
             IF #statPrevOutputValue >= #inputValue
             THEN
               IF #setPosDownRateLim = 0.0
               THEN
                 // set notification for down rate limit in pos range              
                 #tempPosDown := TRUE;
                 IF #inputValue >= 0.0
                 THEN
                   #tempOutv := #inputValue;
                 ELSE
                   #tempOutv := 0.0;
                 END_IF;
               ELSE
                 IF #inputValue >= 0.0
                 THEN
                   // limited rate of change
                   #tempVar := #statPrevOutputValue - #setPosDownRateLim * #tempCycleReal;
                   IF #inputValue < #tempVar
                   THEN
                     // set notification for up rate limit in pos range                  
                     #tempPosDown := TRUE;
                     #tempOutv := #tempVar;
                   END_IF;
                 ELSE  // changeover between pos. and neg. range
                   // period till zero-crossing
                   #tempVar := #statPrevOutputValue / #setPosDownRateLim;

                   IF #tempVar <= #tempCycleReal
                   THEN
                     // limited rate of change
                     #tempVar := - (#tempCycleReal - #tempVar) * #setNegUpRateLim;

                     IF #inputValue < #tempVar
                     THEN
                       // set notification for rate limit
                       #tempPosDown := False;
                       #tempNegUp := TRUE;
                       #tempOutv := #tempVar;
                     END_IF;
                   ELSE
                     // set notification for rate limit
                     #tempPosDown := TRUE;
                     #tempNegUp := FALSE;
                     #tempOutv := #statPrevOutputValue - #tempCycleReal * #setPosDownRateLim;
                   END_IF;
                 END_IF;
               END_IF;
             END_IF;
           END_IF;
         END_IF;
       END_IF;

       // high/low level limitation
       IF #tempOutv >= #setHighLim
       THEN
         #tempHighLim := TRUE;
         IF NOT #statManOp
         THEN
           #tempOutv := #setHighLim;
           // correct up rate limit notification                
           IF #tempOutv - #statPrevOutputValue < #setPosUpRateLim * #tempCycleReal
           THEN
             #tempPosUp := FALSE;
           END_IF;
         END_IF;
       ELSE
         IF #tempOutv <= #setLowLim
         THEN
           #tempLowLim := TRUE;
           IF NOT #statManOp
           THEN
             #tempOutv := #setLowLim;
             // correct up rate limit notification  
             IF #statPrevOutputValue - #tempOutv < #setNegUpRateLim * #tempCycleReal
             THEN
               #tempNegUp := FALSE;
             END_IF;
           END_IF;
         ELSE
           // reset manual mode flag when tempOutv between upper and lower limit        
           #statManOp := FALSE;
         END_IF;
       END_IF;
     END_IF;
   END_IF;


   // update output parameters
   #outputValue := #tempOutv;    // output
   #statPrevOutputValue := #tempOutv;
   #posUpRateLim := #tempPosUp;
   #posDownRateLim := #tempPosDown;
   #negUpRateLim := #tempNegUp;
   #negDownRateLim := #tempNegDown;
   #highLim := #tempHighLim;
   #lowLim := #tempLowLim;
END_FUNCTION_BLOCK

// folder: Phisical_functions/LGF/8 Technology operations/LGF_NonLin

FUNCTION_BLOCK "LGF_NonLin"   // FB10035, SCL
{ S7_Optimized_Access := 'TRUE' }
VERSION : 2.0
   VAR_INPUT
      inputValue : Real;   // Input value
      defaultOutValue : Real;   // Default output value
      onDefaultOutValue : Bool;   // Default output ON: outputValue = defaultOutputValue
      track : Bool;   // Tracking output ON: outputValue = inputValue
      reset : Bool;   // Complete Restart of function block (outputValue = 0.0)
   END_VAR
   VAR_OUTPUT
      outputValue : Real;   // Output value
   END_VAR
   VAR_IN_OUT
      setpoints : Array[*] of "LGF_typeNonLinSetpoints";   // Setpoint table of polynom
   END_VAR
   VAR
      statIndex : Int;   // Index of setpoint table
   END_VAR
   VAR_TEMP
      tempEndOfSearch : Bool;   // End of search algorithm
      tempInputValueStart : Real;   // Actual setpoint - Input value - Low level
      tempInputValueEnd : Real;   // Actual setpoint - Input value - High level
      tempOutputValueStart : Real;   // Actual setpoint - Output value - Low level
      tempOutputValueEnd : Real;   // Actual setpoint - Output value - High level
      tempFactor : Real;   // Gradient of the straight line
      tempLowerBound : Int;   // -
      tempUpperBound : Int;   // -
   END_VAR
BEGIN
   //=============================================================================
   // SIEMENS AG
   // (c)Copyright 2017
   //-----------------------------------------------------------------------------
   // Library:      LGF(Library General Functions)
   // System:       CPU1212C DC/DC/DC FW:V4.2
   // Engineering:  TIA Portal V14 Update 1
   // Restrictions: -
   // Requirements: PLC (S7-1200 FW: 4.2 / S7-1500 FW: 2.0) or higher
   //-----------------------------------------------------------------------------
   // Change log table:
   // Version date         In charge / Changes applied
   // 01.00.00 04.01.2017  Siemens Industry Online Support
   //                      First released version
   // 01.00.01 17.08.2018  Siemens Industry Online Support
   //                      Upgrade: TIA V15 Update 2
   // 01.00.02 23.11.2018  Siemens Industry Online Support
   //                      Upgrade: TIA V15.1
   //=============================================================================

   //Call "LOWER_BOUND" and "UPPER_BOUND" for the setpoints
   #tempLowerBound := DINT_TO_INT(LOWER_BOUND(ARR := #setpoints, DIM := 1));
   #tempUpperBound := DINT_TO_INT(UPPER_BOUND(ARR := #setpoints, DIM := 1));

   //Check index value
   IF (#statIndex < #tempLowerBound) OR (#statIndex > #tempUpperBound) OR (#statIndex = 0)
   THEN
     #statIndex := #tempLowerBound + 1;
   END_IF;

   //Mode: complete restart
   IF (#reset = True)
   THEN
     //Preset search index of array
     #statIndex := #tempLowerBound + 1;
     #outputValue := 0.0;
   ELSE
     //Mode: tracking output
     IF (#track = True)
     THEN
       //Set output value
       #outputValue := #inputValue;
     ELSE
       //Mode: calculated polynom output
       //Initialize search procedure
       #tempEndOfSearch := False;
       //Search procedure
       REPEAT
         //Preset input values of polygon
         #tempInputValueStart := #setpoints[#statIndex - 1].InputValue;
         #tempInputValueEnd := #setpoints[#statIndex].InputValue;
         //Check actual polynom
         IF (#inputValue > #tempInputValueStart)
         THEN
           IF (#inputValue > #tempInputValueEnd)
           THEN
             IF (#statIndex < #tempUpperBound)
             THEN
               #tempInputValueStart := #tempInputValueEnd;
               #statIndex := #statIndex + 1;
               #tempInputValueEnd := #setpoints[#statIndex].InputValue;
             ELSE
               #tempEndOfSearch := True;
             END_IF;
           ELSE
             #tempEndOfSearch := True;
           END_IF;
         ELSE
           IF (#statIndex > (#tempLowerBound + 1))
           THEN
             #statIndex := #statIndex - 1;
             #tempInputValueEnd := #tempInputValueStart;
             // #tempInputValueStart := #setpoints.Point[#statIndex - 1].InputValue;
             #tempInputValueStart := #setpoints[#statIndex].InputValue;
           ELSE
             #tempEndOfSearch := True;
           END_IF;
         END_IF;
       UNTIL
         (#tempEndOfSearch = True)
       END_REPEAT;
       //Set output values of polygon
       #tempOutputValueStart := #setpoints[#statIndex - 1].OutputValue;
       #tempOutputValueEnd := #setpoints[#statIndex].OutputValue;
       //Calculate gradient of straight line
       #tempFactor := (#tempOutputValueEnd - #tempOutputValueStart) / (#tempInputValueEnd - #tempInputValueStart);
       //Calculate output value
       #outputValue := (#tempFactor * #inputValue) + (#tempOutputValueStart - (#tempFactor * #tempInputValueStart));
     END_IF;
   END_IF;

   //Mode: default output
   IF (#onDefaultOutValue = True)
   THEN
     //Set output value
     #outputValue := #defaultOutValue;
   END_IF;
END_FUNCTION_BLOCK

// folder: Phisical_functions/LGF/8 Technology operations/LGF_Ramp

FUNCTION_BLOCK "LGF_Ramp"   // FB10034, SCL
{ S7_Optimized_Access := 'TRUE' }
VERSION : 0.1
   VAR_INPUT
      defaultOutValue : Real := 0.0;   // Default value for preset output
      contStepNbr : Int := 0;   // Hold: continue step number
      contStepTime : Time := T#0MS;   // Hold: time till continue step number
      onDefaulftOutValue : Bool := FALSE;   // Preset output by default value
      start : Bool := FALSE;   // Start operating the timetable
      hold : Bool := FALSE;   // Freeze output at actual value
      continue : Bool := FALSE;   // Hold: prepair continue conditions
      cyclicOP : Bool := FALSE;   // Cyclic timetable operation
      updateTime : Bool := FALSE;   // Update time
      reset : Bool := FALSE;   // Complete reset
      callOB : OB_Cyclic;   // Call OB
   END_VAR
   VAR_OUTPUT
      outputValue : Real;   // Output
      actTimeTable : Bool;   // Time table operation active
      stepNumber : Int;   // Actual step number
      remainTime : Time;   // Remaining time till actual step
      totalTime : Time;   // Total time for time table
      remainTotalTime : Time;   // Remaining total time
      error : Bool;   // -
      statusID : UInt;   // -
      status : Word;   // -
   END_VAR
   VAR_IN_OUT
      setpoints : Array[*] of "LGF_typeRampTimeTable";   // Setpoints for the curve
   END_VAR
   VAR
      statEndValue : Real;   // -
      statOldValue : Real := 0.0;   // -
      statActualStep : Int;   // -
      statActualRestTime : Time;   // -
      statTotalTime : Time;   // -
      statRestTotalTime : Time;   // -
      statStart : Bool;   // -
      statTimeTableActiv : Bool;   // -
      statStartMem : Bool;   // -
      statUpdateTime : Bool;   // -
      statReset : Bool;   // -
      statResetMem : Bool;   // -
   END_VAR
   VAR_TEMP
      tempNewValue : Real;   // -
      tempCounter : Int;   // -
      tempArrayLowLim : DInt;   // -
      tempArrayUpLim : DInt;   // -
      tempReadTimeStatus : Int;   // -
      tempSampleTime : Time;   // -
      tempCycleTime : UDInt;   // -
      tempCyclePhase : UDInt;   // -
      tempCycleStatus : Word;   // -
      tempStart : Bool;   // -
      tempUpdateTime : Bool;   // -
      tempReset : Bool;   // -
   END_VAR
   VAR CONSTANT
      ERROR_QRY_CINT : UInt := 2;   // Error in the instruction "QRY_CINT"
      ERROR_IN_THIS_BLOCK : UInt := 1;   // Error in this block
      NO_ERROR : Word := 16#0000;   // No errors, job finished
      INITIAL : Word := 16#7000;   // Initial values
      FIRST_CALL : Word := 16#7001;   // First call
      FURTHER_CALLS : Word := 16#7002;   // Further calls, cyclic operation
      OB_UNAVAILABLE : Word := 16#8200;   // Call OB unavailable
      ARRAY_LOWER_BOUND : Word := 16#8201;   // Array does not start with 0
   END_VAR
BEGIN
   //=============================================================================
   // Siemens AG
   // (c)Copyright 2017
   //-----------------------------------------------------------------------------
   // Library:       LGF (Library General Functions) 
   // Tested with:   CPU1212C DC/DC/DC FW:V4.2
   // Engineering:   TIA Portal V14 Update 1 
   // Restrictions:  callable only in cyclic interrupt OB
   // Requirements:  PLC (S7-1200 FW: 4.2 / S7-1500 FW: 2.0) or higher
   // Functionality: This function interpolates between defined setpoints.
   //-----------------------------------------------------------------------------
   // Change log table:
   // Version  Date        In charge / Changes applied
   // 01.00.00 03.02.2017  Siemens Industry Online Support
   //                      First released version
   // 01.00.01 16.05.2017  Siemens Industry Online Support
   //                      Comment correction (REGION)
   // 01.00.02 17.08.2018  Siemens Industry Online Support
   //                      Upgrade: TIA V15 Update 2
   // 01.00.03 23.11.2018  Siemens Industry Online Support
   //                      Upgrade: TIA V15.1
   //-----------------------------------------------------------------------------
   //Status Codes:
   // 16#0000:  No errors, job finished
   // 16#7000:  Initial values
   // 16#7001:  First call
   // 16#7002:  Further calls, cyclic operation
   // 16#8200:  Call OB unavailable
   // 16#8201:  Array does not start with 0
   //=============================================================================

   //***// no error
   #error := FALSE;
   #statusID := #ERROR_IN_THIS_BLOCK;

   REGION Cycle time
     //***// get sample time, according to the cyclic interrupt OB number
     #tempReadTimeStatus := QRY_CINT(OB_NR := #callOB, CYCLE => #tempCycleTime, PHASE => #tempCyclePhase, STATUS => #tempCycleStatus);
     #tempCycleTime := #tempCycleTime / 1000; // microsecond --> milisecond 
     #tempSampleTime := UDINT_TO_TIME(#tempCycleTime); // Format: TIME

     // Generate error message of the QRY_CINT function
     IF (#tempReadTimeStatus <> 0) THEN
       #error := TRUE;
       #statusID := #ERROR_QRY_CINT;
       #status := INT_TO_WORD(#tempReadTimeStatus);
       RETURN;
     END_IF;

     // Generate error message when OB unavailable
     IF #tempCycleStatus = 16#0000 THEN
       #error := TRUE;
       #statusID := #ERROR_IN_THIS_BLOCK;
       #status := #OB_UNAVAILABLE;
       RETURN;
     END_IF;
   END_REGION // Cycle time

   REGION Array lower/upper bound
     #tempArrayLowLim := LOWER_BOUND(ARR := #setpoints, DIM := 1);
     #tempArrayUpLim := UPPER_BOUND(ARR := #setpoints, DIM := 1);

     IF #tempArrayLowLim <> 0 THEN
       #error := TRUE;
       #statusID := #ERROR_IN_THIS_BLOCK;
       #status := #ARRAY_LOWER_BOUND;
       RETURN;
     END_IF;
   END_REGION // Array lower/upper bound

   REGION Function 
     #tempUpdateTime := #updateTime AND NOT #statUpdateTime;
     #statUpdateTime := #updateTime;

     REGION First Call
       #tempStart := #start AND NOT #statStartMem;
       #statStartMem := #start;

       IF #tempStart THEN
         #status := #FIRST_CALL;
         #statStart := TRUE;
         #statTotalTime := T#0s;      // reset total time 

         FOR #tempCounter := #tempArrayLowLim TO #tempArrayUpLim // calculate total time 
         DO
           #statTotalTime := #statTotalTime + #setpoints[#tempCounter]."time"; // total time 
         END_FOR;
         #statRestTotalTime := #statTotalTime;
         #statReset := FALSE;
       END_IF;
     END_REGION // First Call

     REGION Reset
       #tempReset := #reset AND NOT #statResetMem;
       #statResetMem := #reset;

       IF #tempReset
       THEN
         //***// RESET 
         #status := #INITIAL;
         #statTotalTime := T#0s;      // reset total time 

         FOR #tempCounter := #tempArrayLowLim TO #tempArrayUpLim // calculate total time 
         DO
           #statTotalTime := #statTotalTime + #setpoints[#tempCounter]."time"; // total time 
         END_FOR;

         #tempNewValue := 0.0;                   // output outValue = 0 
         #statRestTotalTime := #statTotalTime;   // update remaining total time 
         #statEndValue := 0.0;                   // reset statEndValue    
         #statActualStep := 0;                   // reset statActualStep  
         #statActualRestTime := T#0s;            // reset statActualTime 
         #statStart := TRUE;                     // set start condition 
         #statTimeTableActiv := FALSE;           // reset statTimeTableActive 
         #statReset := TRUE;
       END_IF;
     END_REGION // Reset

     REGION Operation 
       IF #start AND NOT #statReset
       THEN
         //***// start function ramp soak 
         IF #statStart
         THEN
           //***// Set up start conditions 
           #tempNewValue := #setpoints[#tempArrayLowLim].outVal;
           #statEndValue := #setpoints[#tempArrayLowLim + 1].outVal;
           #statActualRestTime := #setpoints[#tempArrayLowLim]."time";
           #statRestTotalTime := #statTotalTime;
           #statActualStep := 1;
           #statStart := FALSE;
           #statTimeTableActiv := TRUE;
         ELSE
           IF #hold
           THEN
             //***// Freeze operation 
             #statTimeTableActiv := FALSE;
             #tempNewValue := #statOldValue;

             IF #continue
             THEN
               //***// Set up continue conditions 

               //***// Continue step and remaining time untill continue step
               #statEndValue := #setpoints[#contStepNbr].outVal;
               #statRestTotalTime := #contStepTime;
               #statActualRestTime := #contStepTime;
               #statActualStep := #contStepNbr;

               FOR #tempCounter := #statActualStep TO #tempArrayUpLim // calculating remaining total time  
               DO
                 #statRestTotalTime := #statRestTotalTime + #setpoints[#tempCounter]."time"; // Remaining total time
               END_FOR;
             END_IF;
           ELSE
             //***// normal operation 

             IF #statActualRestTime > #tempSampleTime    // remaining time until actual step 
             THEN
               //***// calculate new output value, if remaining time has not yet expired
               #tempNewValue := #statOldValue + (#statEndValue - #statOldValue) / DINT_TO_REAL(TIME_TO_DINT(#statActualRestTime)) * UDINT_TO_REAL(#tempCycleTime);
               //***// update remaining time till actual step 
               #statActualRestTime := #statActualRestTime - #tempSampleTime;
               //***// update remaining total time 
               #statRestTotalTime := #statRestTotalTime - #tempSampleTime;
             ELSE
               #statActualRestTime := T#0s;
               //***// remaining actual rest time expired 
               IF #statActualStep < #tempArrayUpLim
               THEN
                 //***// End of step numbers not reached yet    
                 //***// set new end value 
                 #statEndValue := #setpoints[#statActualStep + 1].outVal;
                 //***// set new output value 
                 #tempNewValue := #setpoints[#statActualStep].outVal;
                 //***// new remaining actual time 
                 #statActualRestTime := #setpoints[#statActualStep]."time";
                 #statActualStep := #statActualStep + 1;
                 #statTimeTableActiv := TRUE;
                 #statRestTotalTime := #statRestTotalTime - #tempSampleTime;
               ELSE
                 //***// end of step numbers reached 
                 #status := #NO_ERROR;
                 #statRestTotalTime := T#0s;
                 IF #cyclicOP
                 THEN
                   //***// cyclic operation 
                   #statStart := TRUE;
                   #status := #FURTHER_CALLS;
                 ELSE
                   #statTimeTableActiv := FALSE;
                 END_IF;
                 //***// set new output value 
                 #tempNewValue := #setpoints[#statActualStep].outVal;
               END_IF;
             END_IF;
           END_IF;
         END_IF;
       ELSE
         //***// start not active 
         //***// set start flag, for start preparation 
         //#statStart := TRUE;
         #tempNewValue := 0.0;
         //***//  time table not active 
         #statTimeTableActiv := FALSE;
       END_IF;
     END_REGION // Operation 

     REGION Update time
       //***// Update total time and remaining total time 
       IF #updateTime
       THEN
         #statTotalTime := T#0s;     // reset total time 
         #statRestTotalTime := #statActualRestTime;  // copy remaining actual time to remaining total time

         FOR #tempCounter := #tempArrayLowLim TO #tempArrayUpLim // calculate totel time 
         DO
           #statTotalTime := #statTotalTime + #setpoints[#tempCounter]."time"; // total time 
         END_FOR;

         FOR #tempCounter := #statActualStep TO #tempArrayUpLim // calculate remaining total time 
         DO
           #statRestTotalTime := #statRestTotalTime + #setpoints[#tempCounter]."time";// remaining total time 
         END_FOR;
       END_IF;
       //END_IF;
     END_REGION // Update time

     REGION Default output
       //***// default value activated: overwrite output by default value
       IF #onDefaulftOutValue
       THEN
         #tempNewValue := #defaultOutValue;   // preset output 
         #statTimeTableActiv := FALSE; // timetable not active 
       END_IF;
     END_REGION Default output
   END_REGION // Function 

   REGION Write outputs
     //***// update output parameters 
     #outputValue := #tempNewValue;     // output 
     #statOldValue := #tempNewValue;    // store prvious value 
     #actTimeTable := #statTimeTableActiv;  //time table active 
     #stepNumber := #statActualStep; // number of acting step 
     #remainTime := #statActualRestTime;   // remaining time till actual step 
     #totalTime := #statTotalTime;     // total time 
     #remainTotalTime := #statRestTotalTime;    //remaining total time 
   END_REGION // Write outputs
END_FUNCTION_BLOCK

// folder: Phisical_functions/LGF/9 Measurement operations

FUNCTION_BLOCK "LGF_SimpleSmoothingFB"   // FB2, SCL
TITLE = Enable Template
{ S7_Optimized_Access := 'TRUE' }
AUTHOR : (author)
FAMILY : (family)
VERSION : 1.0
// Template for an FB with Enable / Valid Handling according to PLC Open "Function Blocks for Motion Control" V2.0
   VAR_INPUT
      enable : Bool;   // TRUE: Enable functionality of FB; 0: Disable
      insert : Bool;   // Positive edge inserts a new value
      value : Real;   // The value
   END_VAR
   VAR_OUTPUT
      smoothedValue : Real;   // The smoothed value
      busy : Bool;   // TRUE: FB is working and new output values can be expected
      valid : Bool;   // TRUE: Valid set of outputs available at the FB
      error : Bool;   // Rising edge informs that an error occurred during the execution of
      status : Word := 16#7000;   // Current status of FB
   END_VAR
   VAR
      statErrorUserCleared : Bool;   // Error occured that can only be solved by user; rising edge at enable input necessary
      statErrorAutoCleared : Bool;   // Error occured that can be acknowledged by FB
      statEnableOld : Bool;   // Old value of enable for edge detection
      statValues : Array[0..2] of Real;   // Static array values
      statCount : Int;   // Static value for count
      statInsertOld : Bool;   // Static value for insert
      statNoValues : Bool;   // Static value for no values
   END_VAR
   VAR CONSTANT
      STATUS_NO_CALL : Word := 16#7000;   // Status: No call of FB
      STATUS_FIRST_CALL : Word := 16#7001;   // Status: First call of FB after enabling
      STATUS_SUBSEQUENT_CALL : Word := 16#7002;   // Status: Subsequent call of FB
      STATUS_NOT_ENOUGH_VALUES : Word := 16#9000;   // Status: Not enough values (3 values needed)
   END_VAR
BEGIN
   //=============================================================================
   // SIEMENS AG
   // (c)Copyright 2018
   //-----------------------------------------------------------------------------
   // Library:       LGF (Library General Functions)
   // Tested with:   CPU1212C DC/DC/DC FW:V4.2
   // Engineering:   TIA Portal V15.1 
   // Restrictions:  -
   // Requirements:  PLC (S7-1200 / S7-1500)
   // Functionality: This function block calculates the smoothed values 
   //-----------------------------------------------------------------------------
   // Change log table:
   // Version  Date        In charge / Changes applied
   // 01.00.00 23.11.2018  Siemens Industry Online Support
   //                      First released version
   //=============================================================================

   //Check if FB is disabled
   IF NOT #enable
     AND #statEnableOld
   THEN

     //Error outputs are reset with falling edge of enable input
     #statErrorUserCleared := FALSE;
     #statErrorAutoCleared := FALSE;
     #error := FALSE;
     #status := #STATUS_NO_CALL;

     //Enable and busy are reset with falling edge of enable input
     #valid := FALSE;
     #busy := FALSE;

     //Set old value of enable for edge detection and end execution
     #statEnableOld := #enable;
     RETURN;

     //Check if FB is enabled
   ELSIF #enable
     AND NOT #statEnableOld
   THEN
     //reset static values
     #statCount := 0;
     #statValues[0] := 0.0;
     #statValues[1] := 0.0;
     #statValues[2] := 0.0;
     #smoothedValue := 0.0;

     #statNoValues:=true;

     //Busy is set at rising edge of enable input
     #busy := TRUE;
     //Set status for first call
     #status := #STATUS_FIRST_CALL;
     //Set old value of enable for edge detection and end execution
     #statEnableOld := #enable;
     RETURN;

     //Check if user cleared error in FB occurred
   ELSIF #statErrorUserCleared


   THEN
     #busy := FALSE;
     //Set old value of enable for edge detection and end execution
     #statEnableOld := #enable;
     //No set of status necessary, because status already set when error occured
     RETURN;

     //Check if function block is disabled
   ELSIF NOT #enable
   THEN
     #busy := FALSE;
     #status := #STATUS_NO_CALL;
     //Set old value of enable for edge detection and end execution
     #statEnableOld := #enable;
     RETURN;

   ELSE
     //Detect edge for disabling
     #statEnableOld := #enable;
   END_IF;


   //----------------------------------------------------------------------------------------------
   //set Status "Not enough values" after reset
   IF #enable
     AND #statEnableOld
     AND #statNoValues
   THEN
     #status := #STATUS_NOT_ENOUGH_VALUES;
     #statErrorAutoCleared := true;
     #statNoValues := false;
   END_IF;

   // positive edge of insert detected 
   IF #insert
     AND NOT #statInsertOld
   THEN

     #statInsertOld := #insert;
     //copy new value
     #statValues[0] := #statValues[1];
     #statValues[1] := #statValues[2];
     #statValues[2] := #value;

     IF #statCount < 2
     THEN
       #statCount += 1;
       #status := #STATUS_NOT_ENOUGH_VALUES;
       #statErrorAutoCleared := true;
     ELSE
       //3 values inserted, calculate smoothed value
       #smoothedValue := (#statValues[0] + #statValues[1] + #statValues[2]) / 3;
       #statErrorAutoCleared := false;
     END_IF;

   ELSE

     #statInsertOld := #insert;
   END_IF;

   //----------------------------------------------------------------------------------------------
   //Error handling 
   //----------------------------------------------------------------------------------------------
   IF #statErrorUserCleared
   THEN
     #valid := FALSE;
     #busy := FALSE;
     #error := TRUE;

     RETURN;

   ELSIF #statErrorAutoCleared
   THEN
     #valid := FALSE;
     #busy := TRUE;
     #error := TRUE;

     RETURN;

   ELSE
     //Process normal output values
     #valid := TRUE;
     #error := FALSE;
     #status := #STATUS_SUBSEQUENT_CALL; //Set status for subsequent call
   END_IF;
   //----------------------------------------------------------------------------------------------
END_FUNCTION_BLOCK

FUNCTION_BLOCK "LGF_FloatingAverage"   // FB5, SCL
{ S7_Optimized_Access := 'TRUE' }
AUTHOR : SIOS
FAMILY : Math
VERSION : 0.1
   VAR_INPUT
      value : Real;   // Input values REAL
      mode : Int := 1;   // Default mode =1 (triggered); mode= 2 (cyclic)
      windowSize : Int := 100;   // Calculation window of floating average / -
      trigger : Bool;   // Trigger variable
      reset : Bool;   // Trigger for reset
   END_VAR
   VAR_OUTPUT
      average : LReal;   // Floating average
      windowSizeReached : Bool;   // -
      error : Bool;   // "0" = no error; "1" = error
      status : Word;   // status and error codes
   END_VAR
   VAR
      statCounter : Int;   // -
      statTrigger : Bool;   // -
      statValues : Array[0..#MAX_WINDOW_SIZE] of LReal;   // -
      statValuesSum : LReal;   // -
      statWindowSizeOld : Int;   // -
   END_VAR
   VAR_TEMP
      tempTrigger : Bool;   // -
      tempArithmeticAverage : LReal;   // -
      tempCounter : Int;   // -
      tempIndex : Int;
   END_VAR
   VAR CONSTANT
      MAX_WINDOW_SIZE : Int := 100;   // Number of prev. values for floating average
      TRIGGER_MODE : Int := 1;   // Mode: triggered
      CYCLIC_MODE : Int := 2;   // Mode: cyclic
      NO_ERROR : Word := 16#0000;   // -
      NO_MODE : Word := 16#8201;   // Error info: No correct mode selected
      WRONG_WINDOW_SIZE : Word := 16#8202;   // Error info: No correct window size
   END_VAR
BEGIN
   //=============================================================================
   // Siemens AG
   // (c)Copyright 2017
   //-----------------------------------------------------------------------------
   // Library:       LGF (Library General Functions)
   // Tested with:   CPU1212C DC/DC/DC FW:V4.2
   // Engineering:   TIA Portal V14 Update 1
   // Restrictions:  -
   // Requirements:  PLC (S7-1200 / S7-1500)
   // Functionality: This function block calculates the floating arithmetic average
   //                of incoming REAL values each cycle or each trigger impulse.
   //-----------------------------------------------------------------------------
   // Change log table:
   // Version  Date        In charge / Changes applied
   // 01.00.00 16.06.2016  Siemens Industry Online Support
   //                      First released version
   // 01.00.01 02.01.2017  Siemens Industry Online Support
   //                      Upgrade: TIA Portal V14 Update 1
   // 01.01.00 21.02.2017  Siemens Industry Online Support
   //                      Adding variable window size for calculation
   //                      Optimizing calculation algorithm
   // 01.01.01 17.08.2018  Siemens Industry Online Support
   //                      Upgrade: TIA V15 Update 2
   // 01.01.02 23.11.2018  Siemens Industry Online Support
   //                      Upgrade: TIA V15.1
   //-----------------------------------------------------------------------------
   //Status Codes:
   // 16#0000:  No errors
   // 16#8201:  No correct mode selected
   // 16#8202:  No correct window size
   //=============================================================================

   // Set no errors
   #error := FALSE;
   #status := #NO_ERROR;

   // Reset the calculation
   IF #reset THEN
     #average := 0.0;
     #statCounter := 0;
     #statValuesSum := LREAL#0.0;
     #windowSizeReached := FALSE;
     RETURN;
   END_IF;

   // Reset if window size changes
   IF #windowSize <> #statWindowSizeOld THEN
     #average := 0.0;
     #statCounter := 0;
     #statValuesSum := LREAL#0.0;
     #windowSizeReached := FALSE;
     #statWindowSizeOld := #windowSize;
     RETURN;
   END_IF;

   #statWindowSizeOld := #windowSize;

   // Check window size
   IF ((#windowSize > INT#0)
     AND (#windowSize <= #MAX_WINDOW_SIZE)) THEN

     CASE #mode OF // Two modes: Triggered calculation or every cycle
         //--------------------------------------------------------------------------------------------
       #TRIGGER_MODE:
         // This programm code section checks the trigger for a rising edge and sets tempTrigger
         // TRUE in case of a rising edge
         #tempTrigger := #trigger AND NOT #statTrigger;
         #statTrigger := #trigger;

         // Write values into the array #statValues
         IF #tempTrigger THEN // If rising edge of #trigger variable      
           //Calculate array counter
           #tempCounter := #statCounter MOD #windowSize;
           // First filling of the Array with values
           IF (#statCounter < #windowSize) THEN
             //Add value to window
             #tempIndex := #tempCounter;
             #statValues[#tempIndex] := #value;
             //Add value to sum
             #statValuesSum := #statValuesSum + #value;
             //Increment counter
             #statCounter := #statCounter + 1;
             //Calculate avarage value
             #tempArithmeticAverage := #statValuesSum / #statCounter;
           ELSE
             #windowSizeReached := TRUE;
             //Manipulate first value of window
             IF (#tempCounter = INT#0) THEN
               //Add value to sum
               #statValuesSum := #statValuesSum + #value - #statValues[0];
               //Add value to window
               #tempIndex := 0;
               #statValues[#tempIndex] := #value;
               //Increment counter
               #statCounter := #windowSize + 1;
               //Calculate avarage value
               #tempArithmeticAverage := #statValuesSum / #windowSize;
             ELSE
               //Define index
               #tempIndex := #tempCounter;
               //Add value to sum
               #statValuesSum := #statValuesSum + #value - #statValues[#tempIndex];
               //Add value to window
               #statValues[#tempIndex] := #value;
               //Increment counter
               #statCounter := #statCounter + 1;
               //Calculate avarage value
               #tempArithmeticAverage := #statValuesSum / #windowSize;
             END_IF;
           END_IF;

           //Write output
           #average := #tempArithmeticAverage;
         END_IF;
           //--------------------------------------------------------------------------------------------
         #CYCLIC_MODE:
           //Calculate array counter
           #tempCounter := #statCounter MOD #windowSize;
           // First filling of the Array with values
           IF (#statCounter < #windowSize) THEN
             //Add value to window
             #tempIndex := #tempCounter;
             #statValues[#tempIndex] := #value;
             //Add value to sum
             #statValuesSum := #statValuesSum + #value;
             //Increment counter
             #statCounter := #statCounter + 1;
             //Calculate avarage value
             #tempArithmeticAverage := #statValuesSum / #statCounter;
           ELSE
             #windowSizeReached := TRUE;
             //Manipulate first value of window
             IF (#tempCounter = INT#0) THEN
               //Add value to sum
               #statValuesSum := #statValuesSum + #value - #statValues[0];
               //Add value to window
               #tempIndex := 0;
               #statValues[#tempIndex] := #value;
               //Increment counter
               #statCounter := #windowSize + 1;
               //Calculate avarage value
               #tempArithmeticAverage := #statValuesSum / #windowSize;
             ELSE
               //Define index
               #tempIndex := #tempCounter;
               //Add value to sum
               #statValuesSum := #statValuesSum + #value - #statValues[#tempIndex];
               //Add value to window
               #statValues[#tempIndex] := #value;
               //Increment counter
               #statCounter := #statCounter + 1;
               //Calculate avarage value
               #tempArithmeticAverage := #statValuesSum / #windowSize;
             END_IF;
           END_IF;

           //Write output
           #average := #tempArithmeticAverage;
           //--------------------------------------------------------------------------------------------

           // In case of no correct mode was selected setup an error message
         ELSE
           #error := TRUE;
           #status := #NO_MODE; // Info "No correct mode selected"
           #average := 0.0;
           RETURN;
         // END_IF;
     END_CASE;

   ELSE
     // In case of no correct window size setup an error message
     #error := TRUE;
     #status := #WRONG_WINDOW_SIZE; // Info "No correct set of window size"
     #average := 0.0;
   END_IF;
END_FUNCTION_BLOCK

FUNCTION_BLOCK "LGF_Boxplot"   // FB10010, SCL
{ S7_Optimized_Access := 'TRUE' }
VERSION : 0.1
   VAR_INPUT
      execute : Bool;   // Activation of the calculation with each positive edge. / 90.0 degrees
      rangeOutlier : Real := 1.5;   // 0: Outlier detection is deactivated; >1: Outlier detection is activated
   END_VAR
   VAR_OUTPUT
      busy : Bool;   // TRUE: FB is not finished and new output values can be expected
      done : Bool;   // TRUE: Commanded action has been completed successfully
      error : Bool;   // Rising edge informs that an error occurred during the execution of
      status : Word := 16#7000;   // Current status of FB
      statusID : UInt;   // Current statusID of FB
      outlierMax : Real;   // Upper outliers in %.
      max : Real;   // Maximum Value, not an outlier.
      q75 : Real;   // 3rd quartile or Q75 of the data series.
      median : Real;   // 2nd quartile or Median of the data series.
      q25 : Real;   // 1st quartile or Q25 of the data series.
      min : Real;   // Minimum Value, not an outlier.
      outlierMin : Real;   // Lower outliers in %.
      skewness : Real;   // Skewness of the data series.
   END_VAR
   VAR_IN_OUT
      "array" : Variant;   // The data series that is to be used for the calculation
   END_VAR
   VAR
      statMaxNew : Real;   // Static value for Max New
      statMinNew : Real;   // Static value for Min New
      statBusy : Bool;   // Static value for output busy
      statDone : Bool;   // Static value for output done
      statError : Bool;   // Static value for output error
      statExecuteOld : Bool;   // Static value for execute
      instLGF_ShellSortInt : "LGF_ShellSortInt";   // Instance of LG_ShellSortInt
      instLGF_ShellSortReal : "LGF_ShellSortReal";   // Instance of LG_ShellSortReal
      instLGF_ShellSortUInt : "LGF_ShellSortUInt";   // Instance of LG_ShellSortUInt
      statMin : Real;   // Static value for min
      statMax : Real;   // Static value for max
      statQuartil25 : Real;   // Static value for quartil25
      statQuartil75 : Real;   // Static value for quartil75
      statNumberOfElements : UDInt;   // Static value for number of elements
      statEven : Bool;   // Static value for even
      statMedian : Real;   // Static value for median
      statK : Real;   // Static value for K
      statType : Int;   // Static value for type
      statDeltaQuartil : Real;   // Static value for delta quartil
      statOutlierMin : Real;   // Static value for outlier min
      statOutlierMax : Real;   // Static value for outlier max
      statCounter : Int;   // Static value for counter
      statRange : Bool;   // Static value for range
      statBorderOutlier : Real;   // Static value for border outlier
      statRetVal : Int;   // Static value for RetVal
   END_VAR
   VAR_TEMP
      tempValueInt : Int;   // Temporary value for calculation
      tempValueInt1 : Int;   // Temporary value for calculation
      tempValueUint : UInt;   // Temporary value for calculation
      tempValueUint1 : UInt;   // Temporary value for calculation
      tempValueReal : Real;   // Temporary value for calculation
      tempValueReal1 : Real;   // Temporary value for calculation
      tempMinInt : Int;   // Temporary value for min INT
      tempMaxInt : Int;   // Temporary value for max INT
      tempMinUint : UInt;   // Temporary value for min UINT
      tempMaxUint : UInt;   // Temporary value for max UINT
      tempStatus : Word;   // Temporary status
      tempStatusID : UInt;   // Temporary status ID
   END_VAR
   VAR CONSTANT
      OK : Bool := true;   // OK
      NOT_OK : Bool := false;   // NOT_OK
      STATUS_EXECUTION_FINISHED : Word := 16#0000;   // Status: Execution finished without errors
      STATUS_NO_CALL : Word := 16#7000;   // Status: No call of FB
      STATUS_FIRST_CALL : Word := 16#7001;   // Status: First call of FB after enabling
      STATUS_SUBSEQUENT_CALL : Word := 16#7002;   // Status: Subsequent call of FB
      STATUS_RANGE_NOT_OK : Word := 16#9101;   // Status: Range not OK
      STATUS_NO_ARRAY : Word := 16#9102;   // Status: No array
      STATUS_WRONG_DATATYPE : Word := 16#9100;   // Status: Wrong data type
      ID_INTERNAL : UInt := 1;   // Status ID: Internal error
      ID_SORT : UInt := 2;   // Status ID: Error sorting
   END_VAR
BEGIN
   //=============================================================================
   // SIEMENS AG
   // (c)Copyright 2017
   //-----------------------------------------------------------------------------
   // Library:       LGF (Library General Functions)
   // Tested with:   CPU1212C DC/DC/DC FW:V4.2
   // Engineering:   TIA Portal V15.1 
   // Restrictions:  -
   // Requirements:  PLC (S7-1200 / S7-1500)
   // Functionality: The function block sorts the data row and calculates
   //                the so-called "five point summary"
   //-----------------------------------------------------------------------------
   // Change log table:
   // Version  Date        In charge / Changes applied
   // 01.00.00 23.11.2018  Siemens Industry Online Support
   //                      First released version
   //=============================================================================

   //Check if FB is triggered
   IF #execute
     AND NOT #statExecuteOld
     AND NOT #statBusy
   THEN
     //Functionality is busy
     #statBusy := TRUE;
     //#busy := #statBusy;

     //Reset outputs and statics
     #statError := FALSE;
     #status := #STATUS_FIRST_CALL;
     #statDone := FALSE;
     //#done := false;

     #statOutlierMax := 0;
     #statOutlierMin := 0;
     #statMaxNew := 0.0;
     #statMinNew := 0.0;

     #statExecuteOld := #execute;
     GOTO EndOfBlock;
     //FB is currently inactive
   ELSIF NOT #execute
     AND NOT #statBusy
   THEN
     //Error outputs are reset with falling edge of enable input
     #statError := FALSE;

     //Done and busy are reset with falling edge of enable input
     #statDone := FALSE;
     #statBusy := FALSE;

     //Write outputs
     #status := #STATUS_NO_CALL;
     #statExecuteOld := #execute;
     GOTO EndOfBlock;
     //FB is currently executed and not finished
   ELSIF #statBusy
   THEN
     #statExecuteOld := #execute;
     #status := #STATUS_SUBSEQUENT_CALL;
     //FB finished job
   ELSE
     #statExecuteOld := #execute;
     //Wait for start of functionality 
   END_IF;
   //----------------------------------------------------------------------------------------------

   //check RANGE_OUTLIER 
   IF #rangeOutlier = 0
   THEN
     //Value is ok
     #statRange := #OK;
   ELSIF #rangeOutlier <> 0
     AND #rangeOutlier < 1.0
   THEN
     //Value is not ok. Range have to be >1 or 0
     #statRange := #NOT_OK;
     #status := #STATUS_RANGE_NOT_OK;
     #statError := true;
     GOTO EndOfBlock;
   ELSIF #rangeOutlier > 1
   THEN
     //Value is ok
     #statRange := #OK;
   END_IF;


   REGION Program

     //check if input variant is an array
     IF IS_ARRAY(#array)
     THEN
       IF #statError = false
         AND #statBusy = TRUE
         AND #statRange = #OK
       THEN
         //count array elements
         #statNumberOfElements := CountOfElements(#array);

         //check if Number of Elements is even 
         IF (#statNumberOfElements MOD 2) = 0
         THEN
           #statEven := true;
         ELSE
           #statEven := false;
         END_IF;

         //check which datatype is used
         IF TypeOfElements(#array) = Int
         THEN

           REGION Type of array is INT
             //Type is Int
             //Sort array
             #instLGF_ShellSortInt(error => #statError,
                                   statusID => #tempStatusID,
                                   status => #tempStatus,
                                   variantArray := #array);
             IF #statError = true
             THEN
               IF #tempStatusID > 1
               THEN
                 #statusID := #ID_INTERNAL;
               ELSE
                 #statusID := #ID_SORT;
                 #status := #tempStatus;
               END_IF;
               GOTO EndOfBlock;
             ELSE

               //Identify max and min value
               #statRetVal := MOVE_BLK_VARIANT(SRC := #array, COUNT := 1, SRC_INDEX := 0, DEST_INDEX := 0, DEST => #tempMinInt);
               IF #statRetVal <> 0
               THEN
                 #status := INT_TO_WORD(#statRetVal);
                 #statusID := #ID_INTERNAL;
                 #statError := true;
                 GOTO EndOfBlock;
               END_IF;

               #statRetVal := MOVE_BLK_VARIANT(SRC := #array, COUNT := 1, SRC_INDEX := UDINT_TO_INT(#statNumberOfElements - 1), DEST_INDEX := 0, DEST => #tempMaxInt);
               IF #statRetVal <> 0
               THEN
                 #status := INT_TO_WORD(#statRetVal);
                 #statusID := #ID_INTERNAL;
                 #statError := true;
                 GOTO EndOfBlock;
               END_IF;

               #statMax := #tempMaxInt;
               #statMin := #tempMinInt;

               //calculate median (Q50)
               IF #statEven = true
               THEN
                 // if n is even -> calculate MEDIAN = (x(n/2)+x(n/2+1))/2 
                 #statRetVal := MOVE_BLK_VARIANT(SRC := #array, COUNT := 1, SRC_INDEX := UDINT_TO_INT(#statNumberOfElements / 2), DEST_INDEX := 0, DEST => #tempValueInt);
                 IF #statRetVal <> 0
                 THEN
                   #status := INT_TO_WORD(#statRetVal);
                   #statusID := #ID_INTERNAL;
                   #statError := true;
                   GOTO EndOfBlock;
                 END_IF;
                 #statRetVal := MOVE_BLK_VARIANT(SRC := #array, COUNT := 1, SRC_INDEX := UDINT_TO_INT(#statNumberOfElements / 2) - 1, DEST_INDEX := 0, DEST => #tempValueInt1);
                 IF #statRetVal <> 0
                 THEN
                   #status := INT_TO_WORD(#statRetVal);
                   #statusID := #ID_INTERNAL;
                   #statError := true;
                   GOTO EndOfBlock;
                 END_IF;
                 #statMedian := (#tempValueInt1 + #tempValueInt) / 2;
               ELSE
                 // if n is odd -> MEDIAN = x(n+1/2)
                 #statRetVal := MOVE_BLK_VARIANT(SRC := #array, COUNT := 1, SRC_INDEX := UDINT_TO_INT(#statNumberOfElements / 2), DEST_INDEX := 0, DEST => #tempValueInt);
                 IF #statRetVal <> 0
                 THEN
                   #status := INT_TO_WORD(#statRetVal);
                   #statusID := #ID_INTERNAL;
                   #statError := true;
                   GOTO EndOfBlock;
                 END_IF;
                 #statMedian := #tempValueInt;
               END_IF;

               //calculate 1.quartil(Q25)
               // q1 = x(k) with  k=(n+3)/4 
               #statK := (((UDINT_TO_REAL(#statNumberOfElements + 3)) / 4.0)) - 1;
               #statRetVal := MOVE_BLK_VARIANT(SRC := #array, COUNT := 1, SRC_INDEX := TRUNC(#statK), DEST_INDEX := 0, DEST => #tempValueInt);
               IF #statRetVal <> 0
               THEN
                 #status := INT_TO_WORD(#statRetVal);
                 #statusID := #ID_INTERNAL;
                 #statError := true;
                 GOTO EndOfBlock;
               END_IF;
               #statRetVal := MOVE_BLK_VARIANT(SRC := #array, COUNT := 1, SRC_INDEX := TRUNC(#statK) + 1, DEST_INDEX := 0, DEST => #tempValueInt1);
               IF #statRetVal <> 0
               THEN
                 #status := INT_TO_WORD(#statRetVal);
                 #statusID := #ID_INTERNAL;
                 #statError := true;
                 GOTO EndOfBlock;
               END_IF;
               #statQuartil25 := #tempValueInt + FRAC_REAL(#statK) * (#tempValueInt1 - #tempValueInt);

               //calculate 3.quartil(Q75)
               //q3 = x(n+1-k) with k=(3n+1)/4
               #statK := ((3 * UDINT_TO_REAL(#statNumberOfElements) + 1) / 4) - 1;
               #statRetVal := MOVE_BLK_VARIANT(SRC := #array, COUNT := 1, SRC_INDEX := TRUNC(#statK), DEST_INDEX := 0, DEST => #tempValueInt);
               IF #statRetVal <> 0
               THEN
                 #status := INT_TO_WORD(#statRetVal);
                 #statusID := #ID_INTERNAL;
                 #statError := true;
                 GOTO EndOfBlock;
               END_IF;
               #statRetVal := MOVE_BLK_VARIANT(SRC := #array, COUNT := 1, SRC_INDEX := TRUNC(#statK) + 1, DEST_INDEX := 0, DEST => #tempValueInt1);
               IF #statRetVal <> 0
               THEN
                 #status := INT_TO_WORD(#statRetVal);
                 #statusID := #ID_INTERNAL;
                 #statError := true;
                 GOTO EndOfBlock;
               END_IF;
               #statQuartil75 := #tempValueInt + FRAC_REAL(#statK) * (#tempValueInt1 - #tempValueInt);

               //only if RANGE_OUTLIER <> 0
               IF #rangeOutlier <> 0
               THEN

                 //calculate Delta Q75-Q25
                 #statDeltaQuartil := #statQuartil75 - #statQuartil25;

                 //check for min outlier
                 //calculate border for outlier
                 #statBorderOutlier := #statQuartil25 - #rangeOutlier * #statDeltaQuartil;
                 //search in array for values outside the border
                 FOR #statCounter := 0 TO UDINT_TO_INT(#statNumberOfElements - 1) DO
                   #statRetVal := MOVE_BLK_VARIANT(SRC := #array, COUNT := 1, SRC_INDEX := #statCounter, DEST_INDEX := 0, DEST => #tempValueInt);
                   IF #statRetVal <> 0
                   THEN
                     #status := INT_TO_WORD(#statRetVal);
                     #statusID := #ID_INTERNAL;
                     #statError := true;
                     GOTO EndOfBlock;
                   END_IF;
                   IF #tempValueInt < #statBorderOutlier
                   THEN
                     //detected a value as outlier, check next value
                     ;
                   ELSE
                     //all outlier detected. Calulate new Min Value in range and calulate outlier in %
                     #statOutlierMin := INT_TO_REAL((100 * #statCounter)) / UDINT_TO_REAL(#statNumberOfElements);
                     #statMinNew := #tempValueInt;
                     EXIT;
                   END_IF;
                 END_FOR;

